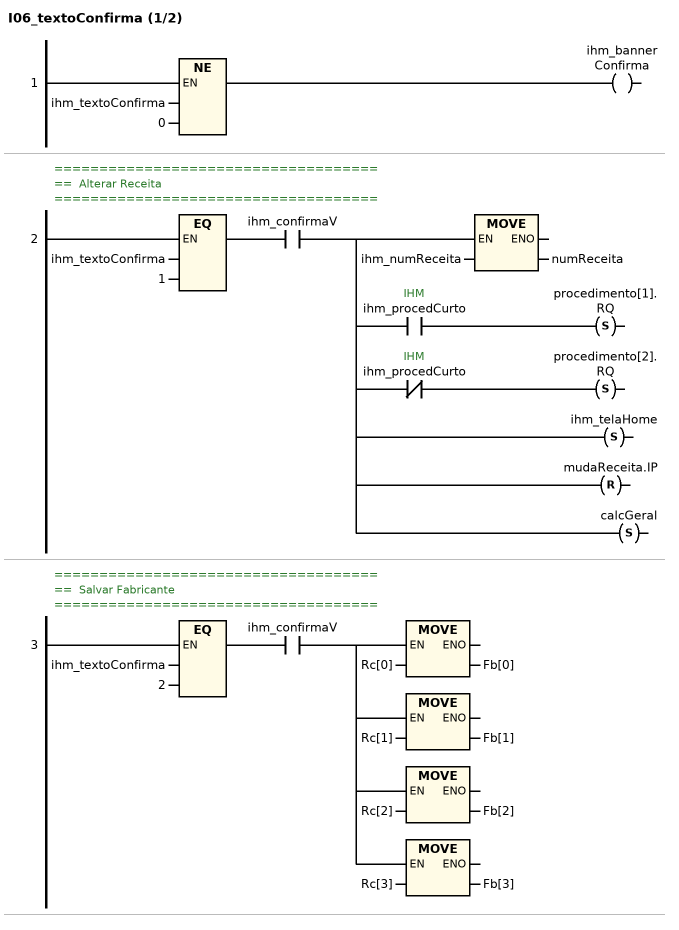
// NETWORK 1
ihm_bannerConfirma := ihm_textoConfirma <> 0;

// NETWORK 2
// ====================================
// ==  Alterar Receita
// ====================================
//   ihm_procedCurto: IHM
_w1 := ihm_textoConfirma = 1 AND ihm_confirmaV;
IF _w1 THEN numReceita := ihm_numReceita; END_IF
procedimento[1].RQ S= _w1 AND ihm_procedCurto;
procedimento[2].RQ S= _w1 AND NOT ihm_procedCurto;
ihm_telaHome S= _w1;
mudaReceita.IP R= _w1;
calcGeral S= _w1;

// NETWORK 3
// ====================================
// ==  Salvar Fabricante
// ====================================
//   Rc[0]: Receita
//   Rc[1]: Receita
//   Rc[2]: Receita
//   Rc[3]: Receita
_w2 := ihm_textoConfirma = 2 AND ihm_confirmaV;
IF _w2 THEN Fb[0] := Rc[0]; END_IF
IF _w2 THEN Fb[1] := Rc[1]; END_IF
IF _w2 THEN Fb[2] := Rc[2]; END_IF
IF _w2 THEN Fb[3] := Rc[3]; END_IF

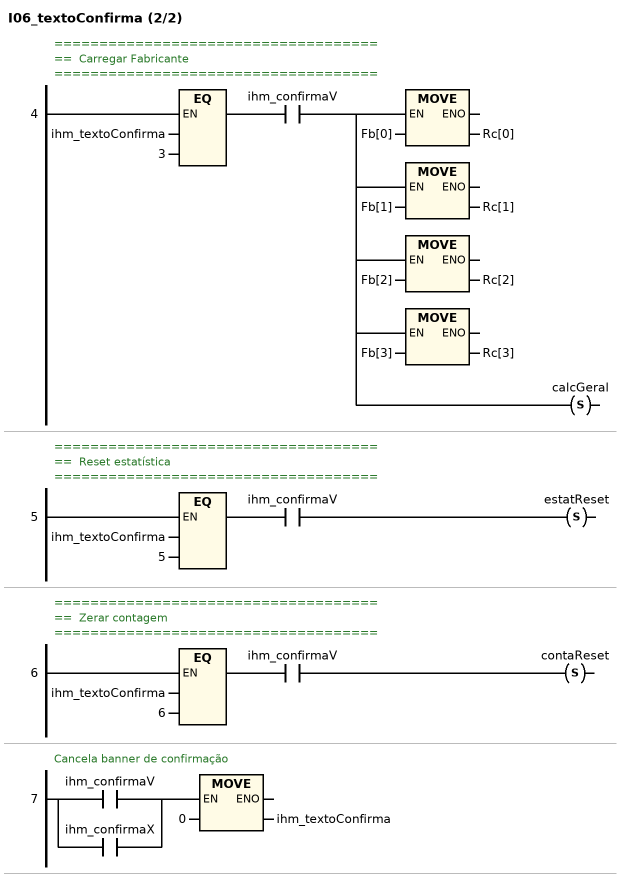
// NETWORK 4
// ====================================
// ==  Carregar Fabricante
// ====================================
//   Rc[0]: Receita
//   Rc[1]: Receita
//   Rc[2]: Receita
//   Rc[3]: Receita
_w3 := ihm_textoConfirma = 3 AND ihm_confirmaV;
IF _w3 THEN Rc[0] := Fb[0]; END_IF
IF _w3 THEN Rc[1] := Fb[1]; END_IF
IF _w3 THEN Rc[2] := Fb[2]; END_IF
IF _w3 THEN Rc[3] := Fb[3]; END_IF
calcGeral S= _w3;

// NETWORK 5
// ====================================
// ==  Reset estatística
// ====================================
estatReset S= ihm_textoConfirma = 5 AND ihm_confirmaV;

// NETWORK 6
// ====================================
// ==  Zerar contagem
// ====================================
contaReset S= ihm_textoConfirma = 6 AND ihm_confirmaV;

// NETWORK 7
// Cancela banner de confirmação
IF ihm_confirmaV OR ihm_confirmaX THEN ihm_textoConfirma := 0; END_IF

END_PROGRAM

// MyController/Application/05_IHM/I07_procedimento
PROGRAM I07_procedimento
VAR
END_VAR
VAR // added by the converter: edge detectors and wires of the graphical bodies
    _w1, _w2, _w3, _w4 : BOOL;
END_VAR

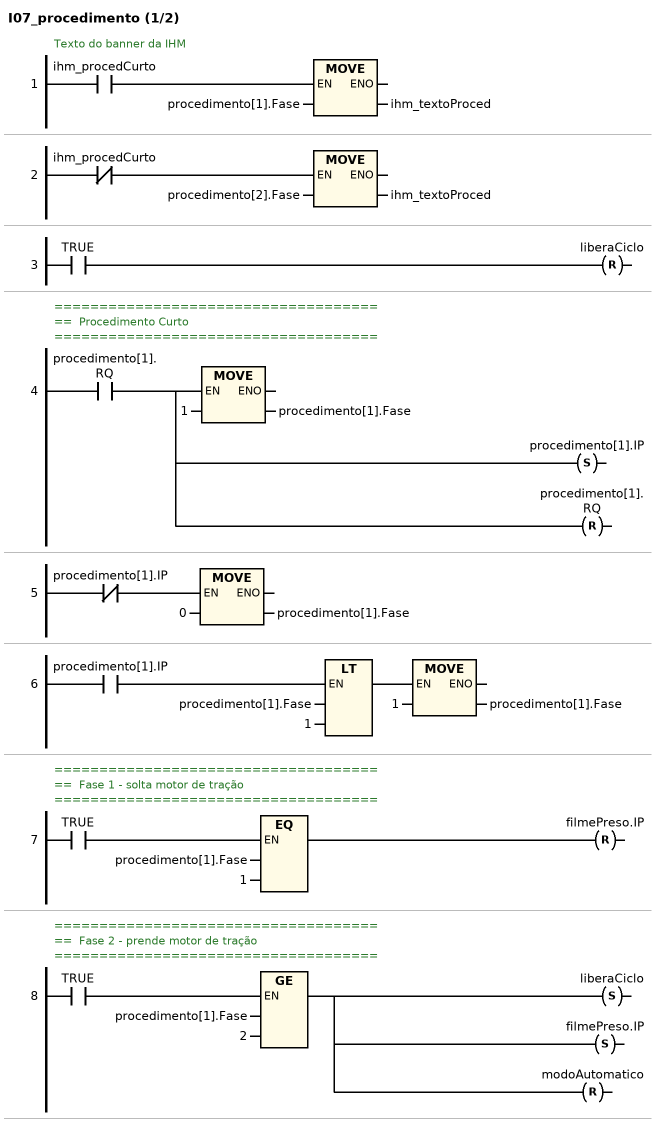
// NETWORK 1
// Texto do banner da IHM
IF ihm_procedCurto THEN ihm_textoProced := procedimento[1].Fase; END_IF

// NETWORK 2
IF NOT ihm_procedCurto THEN ihm_textoProced := procedimento[2].Fase; END_IF

// NETWORK 3
liberaCiclo R= TRUE;

// NETWORK 4
// ====================================
// ==  Procedimento Curto
// ====================================
_w1 := procedimento[1].RQ;
IF _w1 THEN procedimento[1].Fase := 1; END_IF
procedimento[1].IP S= _w1;
procedimento[1].RQ R= _w1;

// NETWORK 5
IF NOT procedimento[1].IP THEN procedimento[1].Fase := 0; END_IF

// NETWORK 6
IF procedimento[1].IP AND procedimento[1].Fase < 1 THEN procedimento[1].Fase := 1; END_IF

// NETWORK 7
// ====================================
// ==  Fase 1 - solta motor de tração
// ====================================
filmePreso.IP R= procedimento[1].Fase = 1;

// NETWORK 8
// ====================================
// ==  Fase 2 - prende motor de tração
// ====================================
_w2 := procedimento[1].Fase >= 2;
liberaCiclo S= _w2;
filmePreso.IP S= _w2;
modoAutomatico R= _w2;

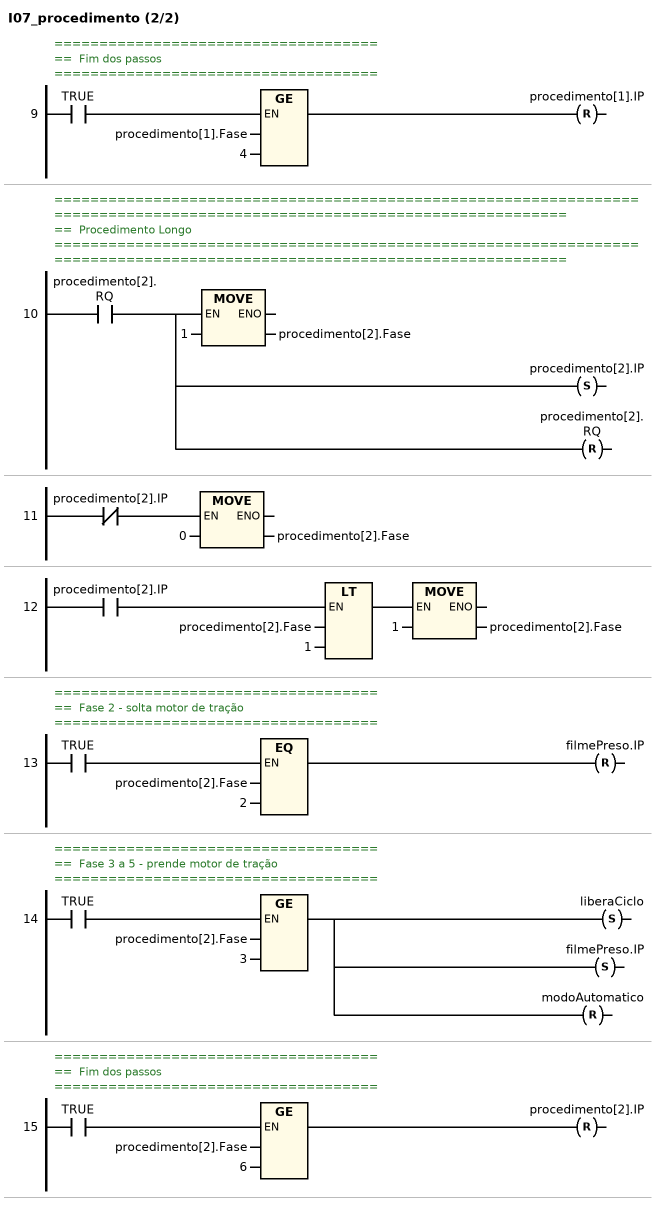
// NETWORK 9
// ====================================
// ==  Fim dos passos
// ====================================
procedimento[1].IP R= procedimento[1].Fase >= 4;

// NETWORK 10
// ==========================================================================================================================
// ==  Procedimento Longo
// ==========================================================================================================================
_w3 := procedimento[2].RQ;
IF _w3 THEN procedimento[2].Fase := 1; END_IF
procedimento[2].IP S= _w3;
procedimento[2].RQ R= _w3;

// NETWORK 11
IF NOT procedimento[2].IP THEN procedimento[2].Fase := 0; END_IF

// NETWORK 12
IF procedimento[2].IP AND procedimento[2].Fase < 1 THEN procedimento[2].Fase := 1; END_IF

// NETWORK 13
// ====================================
// ==  Fase 2 - solta motor de tração
// ====================================
filmePreso.IP R= procedimento[2].Fase = 2;

// NETWORK 14
// ====================================
// ==  Fase 3 a 5 - prende motor de tração
// ====================================
_w4 := procedimento[2].Fase >= 3;
liberaCiclo S= _w4;
filmePreso.IP S= _w4;
modoAutomatico R= _w4;

// NETWORK 15
// ====================================
// ==  Fim dos passos
// ====================================
procedimento[2].IP R= procedimento[2].Fase >= 6;

END_PROGRAM

// MyController/Application/10_Relogio/AjustaDataHora
PROGRAM AjustaDataHora
VAR
	writeDateTime			: SetDateAndTime;
	readDateTime			: GetDateAndTime;
	bitScan					: BOOL;
	comOk					: BOOL;
	T_com					: TON;
END_VAR
VAR // added by the converter: edge detectors and wires of the graphical bodies
    _rt1 : R_TRIG;
END_VAR

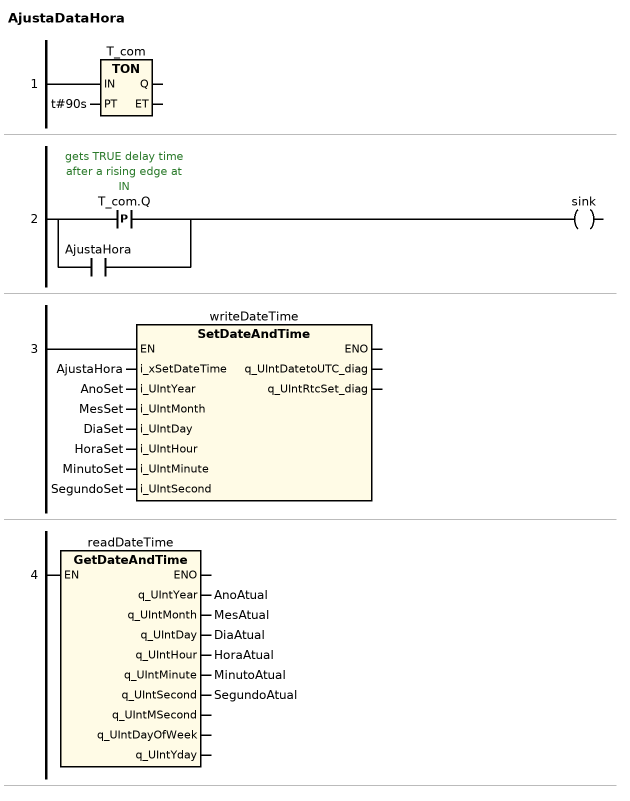
// NETWORK 1
T_com(IN := TRUE, PT := t#90s); // TON

// NETWORK 2
//   T_com.Q: gets TRUE delay time after a rising edge at IN
_rt1(CLK := T_com.Q);
sink := _rt1.Q OR AjustaHora;

// NETWORK 3
//   AnoSet: Sincroniza e ajusta o relógio da IHM
writeDateTime(
    i_xSetDateTime := AjustaHora,
    i_UIntYear := AnoSet,
    i_UIntMonth := MesSet,
    i_UIntDay := DiaSet,
    i_UIntHour := HoraSet,
    i_UIntMinute := MinutoSet,
    i_UIntSecond := SegundoSet); // SetDateAndTime

// NETWORK 4
readDateTime(
    q_UIntYear => AnoAtual,
    q_UIntMonth => MesAtual,
    q_UIntDay => DiaAtual,
    q_UIntHour => HoraAtual,
    q_UIntMinute => MinutoAtual,
    q_UIntSecond => SegundoAtual); // GetDateAndTime

END_PROGRAM

// MyController/Application/10_Relogio/SetDateAndTime
FUNCTION_BLOCK SetDateAndTime
VAR_INPUT
	i_xSetDateTime			: BOOL; (* seta novo horário na transição false para true*)
	i_UIntYear				: UINT:=2011; (*Valor para o ano a ser ajustado*)
	i_UIntMonth				: UINT:=1;(*Valor para o mes a ser ajustado*) 
	i_UIntDay				: UINT:=1;(*Valor para o dia a ser ajustado*) 
	i_UIntHour				: UINT:=0; (*Valor para a hora a ser ajustada*)
	i_UIntMinute			: UINT:=0; (*Valor para o minuto a ser ajustado*)
	i_UIntSecond			: UINT:=0;(*Valor para o segundo a ser ajustado*)
END_VAR
VAR_OUTPUT
	q_UIntDatetoUTC_diag	: UDINT; (*Status quando se =0 ok se <>0 erro nas informações de entrada*)
	q_UIntRtcSet_diag		: UDINT; (*Status quando se =0 ok se <>0 erro nas informações de entrada*)
END_VAR
VAR
	My_UTC					: DWORD; 
	MyDateTime				: SYSTIMEDATE; 
	milesec					: UINT:=0;
	dayOfWeek				: UINT:=1;
	yday					: UINT:=1;
END_VAR
VAR // added by the converter: edge detectors and wires of the graphical bodies
    _s1 : SYSTIMEDATE;
    _w1, _w2 : ANY;
END_VAR

// compose _s1 : SYSTIMEDATE
_s1.wYear := i_UIntYear;
_s1.wMonth := i_UIntMonth;
_s1.wDay := i_UIntDay;
_s1.wHour := i_UIntHour;
_s1.wMinute := i_UIntMinute;
_s1.wSecond := i_UIntSecond;
_s1.wMilliseconds := milesec;
_s1.wDayOfWeek := dayOfWeek;
_s1.wYday := yday;
MyDateTime := _s1;
_w1 := SysTimeRtcConvertDateToUtc(pDate := MyDateTime, pdwTimestampUtc := My_UTC);
q_UIntDatetoUTC_diag := _w1;
IF My_UTC <> 16#FFFFFFFF AND i_xSetDateTime THEN _w2 := SysTimeRtcSet(ulTimestamp := My_UTC); END_IF
q_UIntRtcSet_diag := _w2;
i_xSetDateTime := FALSE;

END_FUNCTION_BLOCK

// MyController/Application/10_Relogio/GetDateAndTime
FUNCTION_BLOCK GetDateAndTime
VAR_INPUT
END_VAR
VAR_OUTPUT
	q_UIntYear			: UINT; 
	q_UIntMonth			: UINT; 
	q_UIntDay			: UINT; 
	q_UIntHour			: UINT; 
	q_UIntMinute		: UINT; 
	q_UIntSecond		: UINT; 
	q_UIntMSecond		: UINT; 
	q_UIntDayOfWeek		: UINT; 
	q_UIntYday			: UINT;
END_VAR
VAR
	Ctrl_DateTime		: SYSTIMEDATE; 
	// SysTimeRtcGet operation diag 
	GetTimeResult		: UDINT; 
// SysTimeRtcConvertUtcToDate operation diag 
	UTCtoDate_diag		: UDINT; 
END_VAR
VAR // added by the converter: edge detectors and wires of the graphical bodies
    _w1, _w2 : ANY;
END_VAR

_w1 := SysTimeRtcGet(pResult := GetTimeResult);
_w2 := SysTimeRtcConvertUtcToDate(dwTimestampUtc := _w1, pDate := Ctrl_DateTime);
UTCtoDate_diag := _w2;
q_UIntYear := Ctrl_DateTime.SYSTIMEDATE;
q_UIntMonth := Ctrl_DateTime.wYear;
q_UIntDay := Ctrl_DateTime.wMonth;
q_UIntHour := Ctrl_DateTime.wDay;
q_UIntMinute := Ctrl_DateTime.wHour;
q_UIntSecond := Ctrl_DateTime.wMinute;
q_UIntMSecond := Ctrl_DateTime.wSecond;
q_UIntDayOfWeek := Ctrl_DateTime.wMilliseconds;
q_UIntYday := Ctrl_DateTime.wDayOfWeek;

END_FUNCTION_BLOCK

// MyController/Application/06_bio/B01_controle
PROGRAM B01_controle
VAR
END_VAR

(*====================================
  ==  Salva Usuario
  ====================================*)
IF digital.loginData THEN
	digital.bioUser[iz]:= digital.login; // Salva Usuario
	digital.bioData[iz]:= DiaAtual; // Salva Data 
	digital.bioHora[iz]:= HoraAtual; // Salva Hora
	digital.bioMin[iz]:= MinutoAtual; // Salva Minuto
	digital.bioGui[iz]:= TRUE; // Lanca Evento
	digital.loginData:= FALSE; // Reseta bit
	iz:= iz + 1; // incrementa ponteiro
END_IF

END_PROGRAM

// MyController/Application/06_bio/B02_data
PROGRAM B02_data
VAR
	ih                : DINT;
	t_backUpBio		  : TON;
END_VAR

(*====================================
  ==  Realiza BackUp e limpa Dados
  ====================================*)
IF iz >= 49 THEN
	ihm_realizaBackup:= TRUE;
END_IF

t_backUpBio(IN:=ihm_realizaBackup, PT:= T#5000MS);

IF t_backUpBio.Q THEN
	 ihm_realizaBackup:= FALSE;
	FOR ih:= 0 TO 49 DO
		 digital.bioUser[ih]:= "";
		 digital.bioData[ih]:= 0;
		 digital.bioHora[ih]:= 0;
		 digital.bioMin[ih]:= 0;
		 digital.bioGui[ih]:= FALSE;
		 iz:= 0;
	END_FOR	
	  ih:= 0;
END_IF

END_PROGRAM

// MyController/Application/07_dados/D01_data
PROGRAM D01_data
VAR
	saveOn					: BOOL;
	backUP					: BOOL;
	dadosReset				: BOOL;
	pf						: INT;
	t_backUp				: TON;
END_VAR

(*====================================
  == Salva dados
  ====================================*)
IF ciclo.IP THEN
	IF (AnoAtual > dados.anoProduzindo) THEN
		limpaDados:= TRUE;
	END_IF
	IF (MesAtual > dados.mesProduzindo) THEN
		ihm_backUpProdutividade:= TRUE;
		IF t_backUp.Q THEN
		limpaDados:= TRUE;
		ihm_backUpProdutividade:= FALSE;
		dados.diaProduzindo:= DiaAtual;
		dados.mesProduzindo:= MesAtual;
		END_IF
	END_IF
END_IF

// Tempo para fazer o BackUp
t_backUp(IN:=ihm_backUpProdutividade, PT:= T#200MS);
				
// Limpa os Dados quando o dia e menor que o dia 
IF dados.diaProduzindo < DiaAtual THEN
	 dadosReset:= TRUE;
	 IF dadosReset THEN
		 ihm_produtMedio:= 0;
	     infoTpoProdHrs:= 0;
	     infoTpoProdMin:= 0;
	     dadosReset:= FALSE;
	     dados.diaProduzindo:= DiaAtual;
	 END_IF
END_IF

// Salva os dados no Arrays
IF ciclo.IP  AND NOT ihm_backUpProdutividade THEN
	 saveOn := TRUE;
	  IF saveON THEN
		 pt:= DiaAtual -1;
	 	 dados.horasProduzidas[pt]:=infoTpoProdHrs;
     	 dados.minProduzidos[pt]:=infoTpoProdMin;
	     dados.produtividade[pt]:=ihm_produtMedio;
	     dados.diaProduzido[pt]:= DiaAtual;
	     dados.pontIhm[pt]:= TRUE;
	     dados.mesProduzindo:= MesAtual;
	     dados.anoProduzindo:= AnoAtual;
	     dados.diaProduzindo:= DiaAtual;	 
	END_IF
 ELSE 
	 saveOn := FALSE;
 END_IF

END_PROGRAM

// MyController/Application/07_dados/D02_clean
PROGRAM D02_clean
VAR
	
	pz 						: DINT;
END_VAR

(*====================================
  == Limpa dados
  ====================================*)
IF limpaDados THEN
	 FOR pz:= 0 TO 30 DO 
		dados.diaProduzido[pz]:= 0;
		dados.horasProduzidas[pz]:= 0;
		dados.minProduzidos[pz]:= 0;
		dados.produtividade[pz]:= 0;
		dados.pontIhm[pz]:= FALSE;
	END_FOR
	limpaDados:= FALSE;
END_IF

END_PROGRAM

// MyController/Application/07_dados/D03_view
PROGRAM D03_view
VAR
	p0						: SINT;
	idxDado   				: DINT;
END_VAR

(*====================================
  == GUI
  ====================================*)
FOR p0:=0 TO 8 DO
	idxDado:= (indPainel * 9) + p0;
	
	IF idxDado > 30 THEN
		RETURN;
	END_IF
	
	// Move  de Datas
	panData[p0]:= dados.diaProduzido[idxDado];
	
	// Move de Produtividade
	panProd[p0]:= dados.produtividade[idxDado];
	
	// Move Hora
	panHora[p0]:= dados.horasProduzidas[idxDado];
	
	// Move Min
	panMin[p0]:= dados.minProduzidos[idxDado];

END_FOR

END_PROGRAM

// MyController/Application/07_dados/D04_controleView
PROGRAM D04_controleView
VAR
	ptr						: ARRAY[0..1] OF R_TRIG;
END_VAR

(*====================================
  ==  Controle GUI
  ====================================*)
ptr[0](CLK:= indSub);
ptr[1](CLK:= indSoma);

	IF ptr[0].Q THEN
		IF indPainel > 0 THEN
			indPainel:=  (indPainel - 1);
		END_IF
	END_IF
 
	IF ptr[1].Q  THEN
		IF indPainel < 3 THEN
			indPainel:=  (indPainel + 1);
		END_IF
	END_IF

END_PROGRAM

// MyController/Application/08_manut/U00_valoresMax
PROGRAM U00_valoresMax
VAR
END_VAR

// Valores Max
util.M_ciclosMax[0]:= 400000;	// Mola Selagem
util.M_ciclosMax[1]:= 800000;	// Mola Desbobinador
util.M_ciclosMax[2]:= 1500000;	// Faca
util.M_ciclosMax[3]:= 400000;	// Mordente Movel
util.M_ciclosMax[4]:= 1000000;	// Mordente Fixo
util.M_ciclosMax[5]:= 2500000;	// Compressor
util.M_ciclosMax[6]:= 1000000;	// Sistema de Corte
util.M_ciclosMax[7]:= 500000;	// Preventiva

END_PROGRAM

// MyController/Application/08_manut/U01_controle
PROGRAM U01_controle
VAR
	p1								: SINT;
	p0								: SINT;
END_VAR

(*====================================
  ==  Vida Util - Compara Valores
  ====================================*)  
IF ciclo.IP THEN
	FOR p0:= 0 TO 7 DO
		IF util.ciclos[p1] >= util.M_ciclosMax[p1] THEN
			util.msg[p1] := TRUE;
		END_IF
		p1:= p1 + 1;
	END_FOR
END_IF

p1:= 0;

END_PROGRAM

// MyController/Application/08_manut/U02_soma
PROGRAM U02_soma
VAR
	p1								: SINT;
	p2								: SINT;
	p0								: SINT;
END_VAR

(*====================================
  ==  Vida Util - Soma
  ====================================*)
IF vidaUtil.RQ THEN
		FOR p0:= 0 TO 7 DO
		IF util.habilita[p1] THEN
			util.ciclos[p1]:= util.ciclos[p1] + 1;
		END_IF
		p1:= p1 + 1;
	END_FOR
	vidaUtil.RQ:= FALSE;
END_IF

p1:= 0;

END_PROGRAM

// MyController/Application/08_manut/U03_reset
PROGRAM U03_reset
VAR
	p1								: SINT;
	p2								: SINT;
	p0								: SINT;
	resetCiclos						: BOOL;
END_VAR

(*====================================
  ==  Vida Util - Reset
  ====================================*)
FOR p0:= 0 TO 7 DO
	IF ihm_resetCiclos[p1] THEN
		util.ciclos[p1] := 0;
		ihm_resetCiclos[p1]:= FALSE;
		util.msg[p1]:= FALSE;
	END_IF
		p1:= p1 + 1;
END_FOR

p1:= 0;

END_PROGRAM

// MyController/Application/08_manut/U04_view
PROGRAM U04_view
VAR
	p1								: SINT;
	p2								: SINT:= 15;
	p0								: SINT;
	msgTimer						: TON;
END_VAR

(*====================================
  ==  Aciona Mensagens
  ====================================*)
msgTimer(IN:= msgPrimeiro,
	  	 PT:= T#2S);
				  
IF msgTimer.Q THEN
	FOR p0:= 0 TO 7 DO
		IF util.msg[p1] AND util.habilita[p1] THEN
			alarme[p2] := TRUE;
		END_IF
		p1:= p1 + 1;
		p2:= p2 + 1;
	END_FOR
	msgPrimeiro:= FALSE;
END_IF

END_PROGRAM

// MyController/Application/02_Filme/F04_foto
PROGRAM F04_foto
VAR
END_VAR
VAR // added by the converter: edge detectors and wires of the graphical bodies
    _rt1 : R_TRIG;
    _w1, _w2 : BOOL;
END_VAR

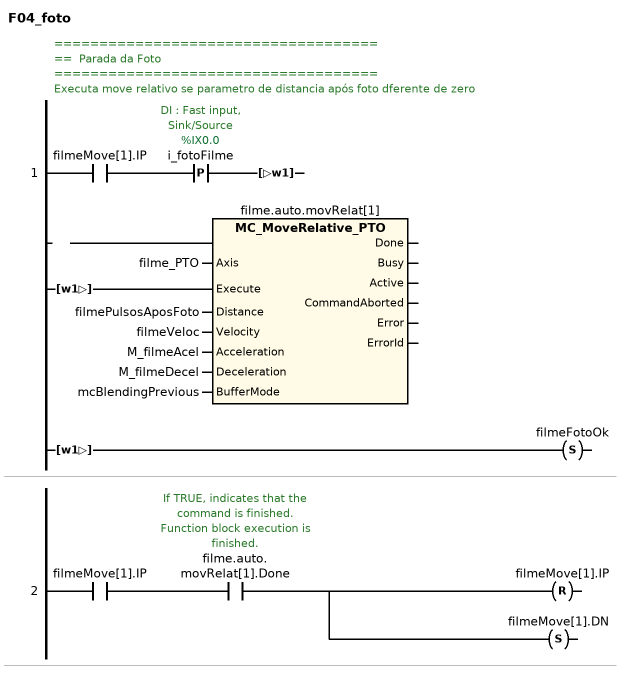
// NETWORK 1
// ====================================
// ==  Parada da Foto
// ====================================
// Executa move relativo se parametro de distancia após foto dferente de zero
//   i_fotoFilme: DI : Fast input, Sink/Source | AT %IX0.0
_rt1(CLK := i_fotoFilme);
_w1 := filmeMove[1].IP AND _rt1.Q;
filme.auto.movRelat[1](
    Axis := filme_PTO,
    Execute := _w1,
    Distance := filmePulsosAposFoto,
    Velocity := filmeVeloc,
    Acceleration := M_filmeAcel,
    Deceleration := M_filmeDecel,
    BufferMode := mcBlendingPrevious); // MC_MoveRelative_PTO
filmeFotoOk S= _w1;

// NETWORK 2
//   filme.auto.movRelat[1].Done: If TRUE, indicates that the command is finished. Function block execution is finished.
_w2 := filmeMove[1].IP AND filme.auto.movRelat[1].Done;
filmeMove[1].IP R= _w2;
filmeMove[1].DN S= _w2;

END_PROGRAM

// MyController/Application/04_Disco/D04_foto
PROGRAM D04_foto
VAR
END_VAR
VAR // added by the converter: edge detectors and wires of the graphical bodies
    _rt1 : R_TRIG;
    _w1 : BOOL;
END_VAR

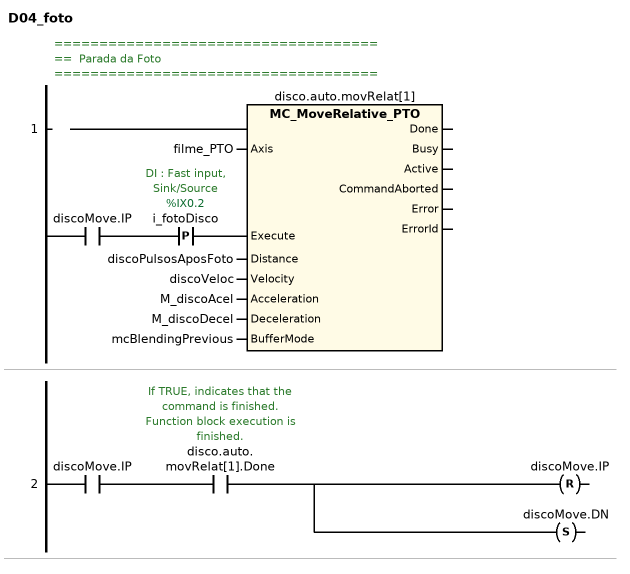
// NETWORK 1
// ====================================
// ==  Parada da Foto
// ====================================
//   i_fotoDisco: DI : Fast input, Sink/Source | AT %IX0.2
_rt1(CLK := i_fotoDisco);
disco.auto.movRelat[1](
    Axis := filme_PTO,
    Execute := discoMove.IP AND _rt1.Q,
    Distance := discoPulsosAposFoto,
    Velocity := discoVeloc,
    Acceleration := M_discoAcel,
    Deceleration := M_discoDecel,
    BufferMode := mcBlendingPrevious); // MC_MoveRelative_PTO

// NETWORK 2
//   disco.auto.movRelat[1].Done: If TRUE, indicates that the command is finished. Function block execution is finished.
_w1 := discoMove.IP AND disco.auto.movRelat[1].Done;
discoMove.IP R= _w1;
discoMove.DN S= _w1;

END_PROGRAM

// MyController/Application/03_Selagem/S06_seguranca
PROGRAM S06_seguranca
VAR
END_VAR
VAR // added by the converter: edge detectors and wires of the graphical bodies
    _ft1 : F_TRIG;
    _w1 : BOOL;
END_VAR

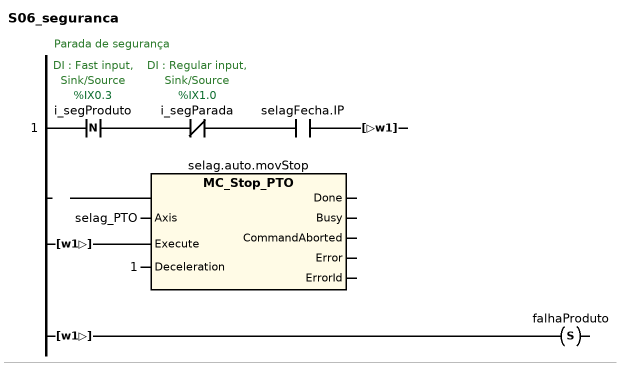
// NETWORK 1
// Parada de segurança
//   i_segProduto: DI : Fast input, Sink/Source | AT %IX0.3
//   i_segParada: DI : Regular input, Sink/Source | AT %IX1.0
_ft1(CLK := i_segProduto);
_w1 := _ft1.Q AND NOT i_segParada AND selagFecha.IP;
selag.auto.movStop(Axis := selag_PTO, Execute := _w1, Deceleration := 1); // MC_Stop_PTO
falhaProduto S= _w1;

END_PROGRAM

// MyController/Application/HiddenPOU
FUNCTION HiddenPOU : BOOL

VAR_INPUT
	pHiddenFunc: POINTER TO WORD;
END_VAR
VAR
	pRead: POINTER TO BYTE;
	pWrite: POINTER TO BYTE;
END_VAR

pRead := pHiddenFunc + 400;
pWrite := pHiddenFunc + 4400;
HiddenPOU := TRUE;

END_FUNCTION

// MyController/Application/Visu/Info
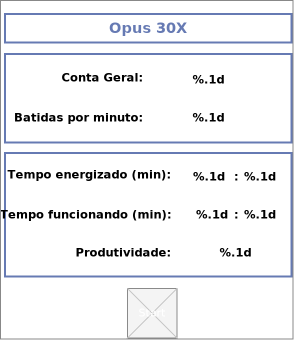
VISUALIZATION Info  // 294x340
    RoundedRectangle (4,152 288x125)
    RoundedRectangle (4,53 288x90)
    Image (127,288 50x50), "Start", image: Imagens.Botao
        OnMouseClick:  ToggleVariable=vsBtStart
    RoundedRectangle (4,13 288x30), "Opus 30X"
    Label (6,60 140x35), "Conta Geral:"
    Label (6,100 140x35), "Batidas por minuto:"
    Rectangle (151,62 115x35), "%.1d", text variable: ihm_contaGeral
    Rectangle (151,100 115x35), "%.1d", text variable: ihm_velocMedida
    Label (4,157 170x35), "Tempo energizado (min):"
    Label (4,197 170x35), "Tempo funcionando (min):"
    Rectangle (173,159 55x35), "%.1d", text variable: infoTpoEnergHrs
    Label (4,235 170x35), "Produtividade:"
    Rectangle (192,235 87x35), "%.1d", text variable: ihm_produtMedio
    Rectangle (241,159 35x35), "%.1d", text variable: infoTpoEnergMin
    Rectangle (176,197 55x35), "%.1d", text variable: infoTpoProdHrs
    Rectangle (241,197 35x35), "%.1d", text variable: infoTpoProdMin
    Label (230,159 13x35), ":"
    Label (230,197 13x35), ":"
END_VISUALIZATION

// MyController/Application/Visu/Main
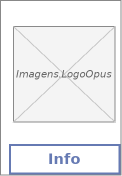
VISUALIZATION Main  // 122x176
    Image (13,26 102x96), image: Imagens.LogoOpus
    RoundedRectangle (9,144 111x30), "Info"
        OnMouseClick:  Assign=Info, Type=Assignment
END_VISUALIZATION
